REGION Network 9: Position Carrier Control First Carrier in Production Zone
   // Control of First Carrier in Zone Closest to end position/Stop.  Move command is issued to carrier. Carrier will move in auto.
   Label( ProdZoneFirstCarrierPosition )
   RUNG wire#powerrail
      Move(in := "EMS".Zone[#Zone].EndPos, out1 => #TrafficCopCarrierZnBufferOut[#CarrierZnArrayPos].CommandPos)
      Sub(in1 := #TrafficCopCarrierZnBufferOut[#CarrierZnArrayPos].CommandPos, in2 := "EMS".Zone[#Zone].InPositionTolerance, out => #TrafficCopCarrierZnBufferOut[#CarrierZnArrayPos].CommandPosLowLimit)
      Add(in1 := #TrafficCopCarrierZnBufferOut[#CarrierZnArrayPos].CommandPos, in2 := "EMS".Zone[#Zone].InPositionTolerance, out => #TrafficCopCarrierZnBufferOut[#CarrierZnArrayPos].CommandPosHighLimit)
   END_RUNG
   RUNG wire#powerrail
      { S7_Templates := "SrcType := DInt" } GE_Contact(in1 := "EMS".Carrier[#CarNumZnPos[1]].Position, in2 := #TrafficCopCarrierZnBufferOut[#CarrierZnArrayPos].CommandPosLowLimit)
      { S7_Templates := "SrcType := DInt" } LE_Contact(in1 := "EMS".Zone[#Zone].EndPos, in2 := #TrafficCopCarrierZnBufferOut[#CarrierZnArrayPos].CommandPosHighLimit)
      Coil( #TrafficCopCarrierZnBufferOut[#CarrierZnArrayPos].AtCommandPos )
   END_RUNG
   RUNG wire#powerrail
      Contact( "EMS".Carrier[#CarNumZnPos[1]].SDC_IN.AutoMode )
      I_Contact( #TrafficCopCarrierZnBufferOut[#CarrierZnArrayPos].AtCommandPos )
      Coil( #TCZnPosnArray.Carrier[#CarNumZnPos[#CarrierZnArrayPos]].MoveFwd )
   END_RUNG
   // the same network as SCL:
   ProdZoneFirstCarrierPosition:
   #TrafficCopCarrierZnBufferOut[#CarrierZnArrayPos].CommandPos := "EMS".Zone[#Zone].EndPos;
   #TrafficCopCarrierZnBufferOut[#CarrierZnArrayPos].CommandPosLowLimit := #TrafficCopCarrierZnBufferOut[#CarrierZnArrayPos].CommandPos - "EMS".Zone[#Zone].InPositionTolerance;
   #TrafficCopCarrierZnBufferOut[#CarrierZnArrayPos].CommandPosHighLimit := #TrafficCopCarrierZnBufferOut[#CarrierZnArrayPos].CommandPos + "EMS".Zone[#Zone].InPositionTolerance;
   #TrafficCopCarrierZnBufferOut[#CarrierZnArrayPos].AtCommandPos := ("EMS".Carrier[#CarNumZnPos[1]].Position >= #TrafficCopCarrierZnBufferOut[#CarrierZnArrayPos].CommandPosLowLimit) AND ("EMS".Zone[#Zone].EndPos <= #TrafficCopCarrierZnBufferOut[#CarrierZnArrayPos].CommandPosHighLimit);
   #TCZnPosnArray.Carrier[#CarNumZnPos[#CarrierZnArrayPos]].MoveFwd := "EMS".Carrier[#CarNumZnPos[1]].SDC_IN.AutoMode AND NOT #TrafficCopCarrierZnBufferOut[#CarrierZnArrayPos].AtCommandPos;
END_REGION

REGION Network 10: Start of 2nd to last Carrier in Zone Carrier Control
   Label( ZoneNextCarrierPosition )
   RUNG wire#powerrail
      Contact( "EMS".Zone[#Zone].AccumZone )
      JumpCoil( AccumZoneNextCarrierPosition )
   END_RUNG
   // the same network as SCL:
   ZoneNextCarrierPosition:
   IF "EMS".Zone[#Zone].AccumZone THEN GOTO AccumZoneNextCarrierPosition; END_IF;
END_REGION

REGION Network 11: Jump to Production Zone 2nd to Last Carrier Position Carrier Control
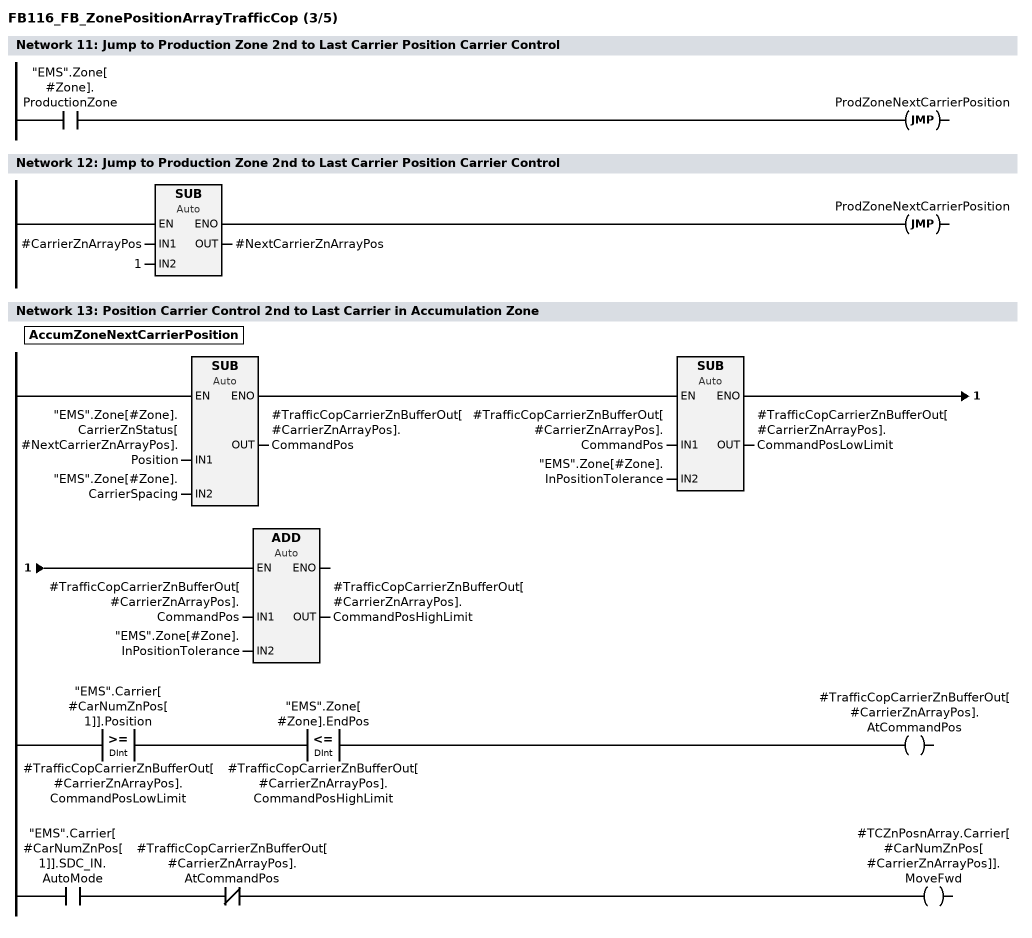
   RUNG wire#powerrail
      Contact( "EMS".Zone[#Zone].ProductionZone )
      JumpCoil( ProdZoneNextCarrierPosition )
   END_RUNG
   // the same network as SCL:
   IF "EMS".Zone[#Zone].ProductionZone THEN GOTO ProdZoneNextCarrierPosition; END_IF;
END_REGION

REGION Network 12: Jump to Production Zone 2nd to Last Carrier Position Carrier Control
   RUNG wire#powerrail
      Sub(in1 := #CarrierZnArrayPos, in2 := 1, out => #NextCarrierZnArrayPos)
      JumpCoil( ProdZoneNextCarrierPosition )
   END_RUNG
   // the same network as SCL:
   #NextCarrierZnArrayPos := #CarrierZnArrayPos - 1;
   GOTO ProdZoneNextCarrierPosition;
END_REGION

REGION Network 13: Position Carrier Control 2nd to Last Carrier in Accumulation Zone
   Label( AccumZoneNextCarrierPosition )
   RUNG wire#powerrail
      Sub(in1 := "EMS".Zone[#Zone].CarrierZnStatus[#NextCarrierZnArrayPos].Position, in2 := "EMS".Zone[#Zone].CarrierSpacing, out => #TrafficCopCarrierZnBufferOut[#CarrierZnArrayPos].CommandPos)
      Sub(in1 := #TrafficCopCarrierZnBufferOut[#CarrierZnArrayPos].CommandPos, in2 := "EMS".Zone[#Zone].InPositionTolerance, out => #TrafficCopCarrierZnBufferOut[#CarrierZnArrayPos].CommandPosLowLimit)
      Add(in1 := #TrafficCopCarrierZnBufferOut[#CarrierZnArrayPos].CommandPos, in2 := "EMS".Zone[#Zone].InPositionTolerance, out => #TrafficCopCarrierZnBufferOut[#CarrierZnArrayPos].CommandPosHighLimit)
   END_RUNG
   RUNG wire#powerrail
      { S7_Templates := "SrcType := DInt" } GE_Contact(in1 := "EMS".Carrier[#CarNumZnPos[1]].Position, in2 := #TrafficCopCarrierZnBufferOut[#CarrierZnArrayPos].CommandPosLowLimit)
      { S7_Templates := "SrcType := DInt" } LE_Contact(in1 := "EMS".Zone[#Zone].EndPos, in2 := #TrafficCopCarrierZnBufferOut[#CarrierZnArrayPos].CommandPosHighLimit)
      Coil( #TrafficCopCarrierZnBufferOut[#CarrierZnArrayPos].AtCommandPos )
   END_RUNG
   RUNG wire#powerrail
      Contact( "EMS".Carrier[#CarNumZnPos[1]].SDC_IN.AutoMode )
      I_Contact( #TrafficCopCarrierZnBufferOut[#CarrierZnArrayPos].AtCommandPos )
      Coil( #TCZnPosnArray.Carrier[#CarNumZnPos[#CarrierZnArrayPos]].MoveFwd )
   END_RUNG
   // the same network as SCL:
   AccumZoneNextCarrierPosition:
   #TrafficCopCarrierZnBufferOut[#CarrierZnArrayPos].CommandPos := "EMS".Zone[#Zone].CarrierZnStatus[#NextCarrierZnArrayPos].Position - "EMS".Zone[#Zone].CarrierSpacing;
   #TrafficCopCarrierZnBufferOut[#CarrierZnArrayPos].CommandPosLowLimit := #TrafficCopCarrierZnBufferOut[#CarrierZnArrayPos].CommandPos - "EMS".Zone[#Zone].InPositionTolerance;
   #TrafficCopCarrierZnBufferOut[#CarrierZnArrayPos].CommandPosHighLimit := #TrafficCopCarrierZnBufferOut[#CarrierZnArrayPos].CommandPos + "EMS".Zone[#Zone].InPositionTolerance;
   #TrafficCopCarrierZnBufferOut[#CarrierZnArrayPos].AtCommandPos := ("EMS".Carrier[#CarNumZnPos[1]].Position >= #TrafficCopCarrierZnBufferOut[#CarrierZnArrayPos].CommandPosLowLimit) AND ("EMS".Zone[#Zone].EndPos <= #TrafficCopCarrierZnBufferOut[#CarrierZnArrayPos].CommandPosHighLimit);
   #TCZnPosnArray.Carrier[#CarNumZnPos[#CarrierZnArrayPos]].MoveFwd := "EMS".Carrier[#CarNumZnPos[1]].SDC_IN.AutoMode AND NOT #TrafficCopCarrierZnBufferOut[#CarrierZnArrayPos].AtCommandPos;
END_REGION

REGION Network 14: Position Carrier Control 2nd to Last Carrier in Production Zone
   // Control of 2nd to Last Carrier in Zone Move to next zone with carrier spacing
   // .  Move command is issued to carrier. Carrier will move in auto.
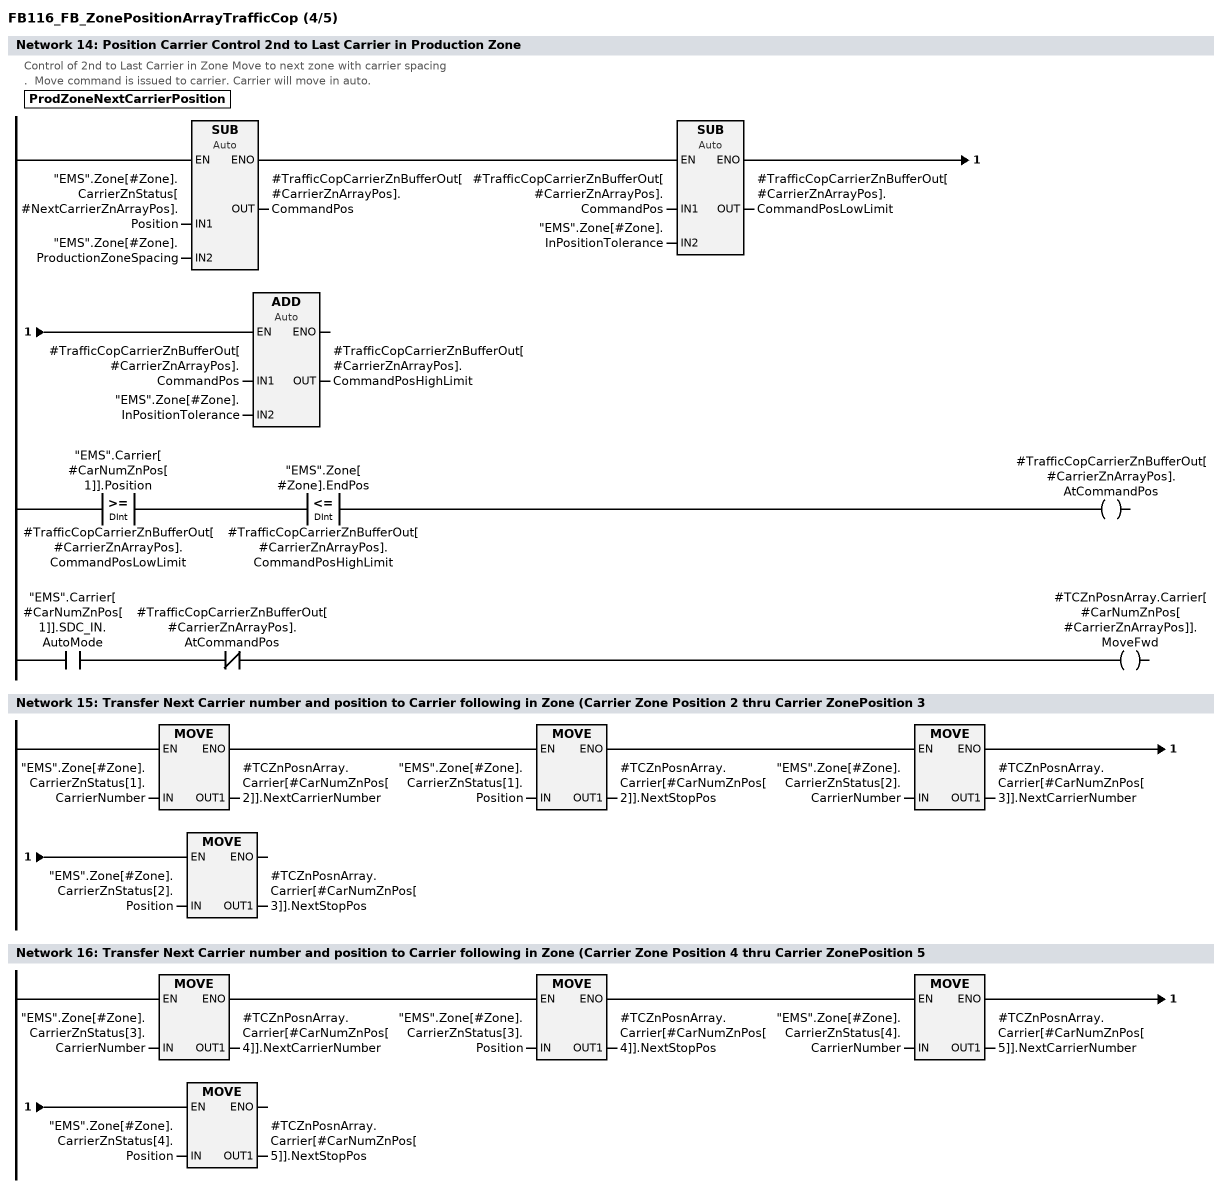
   Label( ProdZoneNextCarrierPosition )
   RUNG wire#powerrail
      Sub(in1 := "EMS".Zone[#Zone].CarrierZnStatus[#NextCarrierZnArrayPos].Position, in2 := "EMS".Zone[#Zone].ProductionZoneSpacing, out => #TrafficCopCarrierZnBufferOut[#CarrierZnArrayPos].CommandPos)
      Sub(in1 := #TrafficCopCarrierZnBufferOut[#CarrierZnArrayPos].CommandPos, in2 := "EMS".Zone[#Zone].InPositionTolerance, out => #TrafficCopCarrierZnBufferOut[#CarrierZnArrayPos].CommandPosLowLimit)
      Add(in1 := #TrafficCopCarrierZnBufferOut[#CarrierZnArrayPos].CommandPos, in2 := "EMS".Zone[#Zone].InPositionTolerance, out => #TrafficCopCarrierZnBufferOut[#CarrierZnArrayPos].CommandPosHighLimit)
   END_RUNG
   RUNG wire#powerrail
      { S7_Templates := "SrcType := DInt" } GE_Contact(in1 := "EMS".Carrier[#CarNumZnPos[1]].Position, in2 := #TrafficCopCarrierZnBufferOut[#CarrierZnArrayPos].CommandPosLowLimit)
      { S7_Templates := "SrcType := DInt" } LE_Contact(in1 := "EMS".Zone[#Zone].EndPos, in2 := #TrafficCopCarrierZnBufferOut[#CarrierZnArrayPos].CommandPosHighLimit)
      Coil( #TrafficCopCarrierZnBufferOut[#CarrierZnArrayPos].AtCommandPos )
   END_RUNG
   RUNG wire#powerrail
      Contact( "EMS".Carrier[#CarNumZnPos[1]].SDC_IN.AutoMode )
      I_Contact( #TrafficCopCarrierZnBufferOut[#CarrierZnArrayPos].AtCommandPos )
      Coil( #TCZnPosnArray.Carrier[#CarNumZnPos[#CarrierZnArrayPos]].MoveFwd )
   END_RUNG
   // the same network as SCL:
   ProdZoneNextCarrierPosition:
   #TrafficCopCarrierZnBufferOut[#CarrierZnArrayPos].CommandPos := "EMS".Zone[#Zone].CarrierZnStatus[#NextCarrierZnArrayPos].Position - "EMS".Zone[#Zone].ProductionZoneSpacing;
   #TrafficCopCarrierZnBufferOut[#CarrierZnArrayPos].CommandPosLowLimit := #TrafficCopCarrierZnBufferOut[#CarrierZnArrayPos].CommandPos - "EMS".Zone[#Zone].InPositionTolerance;
   #TrafficCopCarrierZnBufferOut[#CarrierZnArrayPos].CommandPosHighLimit := #TrafficCopCarrierZnBufferOut[#CarrierZnArrayPos].CommandPos + "EMS".Zone[#Zone].InPositionTolerance;
   #TrafficCopCarrierZnBufferOut[#CarrierZnArrayPos].AtCommandPos := ("EMS".Carrier[#CarNumZnPos[1]].Position >= #TrafficCopCarrierZnBufferOut[#CarrierZnArrayPos].CommandPosLowLimit) AND ("EMS".Zone[#Zone].EndPos <= #TrafficCopCarrierZnBufferOut[#CarrierZnArrayPos].CommandPosHighLimit);
   #TCZnPosnArray.Carrier[#CarNumZnPos[#CarrierZnArrayPos]].MoveFwd := "EMS".Carrier[#CarNumZnPos[1]].SDC_IN.AutoMode AND NOT #TrafficCopCarrierZnBufferOut[#CarrierZnArrayPos].AtCommandPos;
END_REGION

REGION Network 15: Transfer Next Carrier number and position to Carrier following in Zone (Carrier Zone Position 2 thru Carrier ZonePosition 3
   RUNG wire#powerrail
      Move(in := "EMS".Zone[#Zone].CarrierZnStatus[1].CarrierNumber, out1 => #TCZnPosnArray.Carrier[#CarNumZnPos[2]].NextCarrierNumber)
      Move(in := "EMS".Zone[#Zone].CarrierZnStatus[1].Position, out1 => #TCZnPosnArray.Carrier[#CarNumZnPos[2]].NextStopPos)
      Move(in := "EMS".Zone[#Zone].CarrierZnStatus[2].CarrierNumber, out1 => #TCZnPosnArray.Carrier[#CarNumZnPos[3]].NextCarrierNumber)
      Move(in := "EMS".Zone[#Zone].CarrierZnStatus[2].Position, out1 => #TCZnPosnArray.Carrier[#CarNumZnPos[3]].NextStopPos)
   END_RUNG
   // the same network as SCL:
   #TCZnPosnArray.Carrier[#CarNumZnPos[2]].NextCarrierNumber := "EMS".Zone[#Zone].CarrierZnStatus[1].CarrierNumber;
   #TCZnPosnArray.Carrier[#CarNumZnPos[2]].NextStopPos := "EMS".Zone[#Zone].CarrierZnStatus[1].Position;
   #TCZnPosnArray.Carrier[#CarNumZnPos[3]].NextCarrierNumber := "EMS".Zone[#Zone].CarrierZnStatus[2].CarrierNumber;
   #TCZnPosnArray.Carrier[#CarNumZnPos[3]].NextStopPos := "EMS".Zone[#Zone].CarrierZnStatus[2].Position;
END_REGION

REGION Network 16: Transfer Next Carrier number and position to Carrier following in Zone (Carrier Zone Position 4 thru Carrier ZonePosition 5
   RUNG wire#powerrail
      Move(in := "EMS".Zone[#Zone].CarrierZnStatus[3].CarrierNumber, out1 => #TCZnPosnArray.Carrier[#CarNumZnPos[4]].NextCarrierNumber)
      Move(in := "EMS".Zone[#Zone].CarrierZnStatus[3].Position, out1 => #TCZnPosnArray.Carrier[#CarNumZnPos[4]].NextStopPos)
      Move(in := "EMS".Zone[#Zone].CarrierZnStatus[4].CarrierNumber, out1 => #TCZnPosnArray.Carrier[#CarNumZnPos[5]].NextCarrierNumber)
      Move(in := "EMS".Zone[#Zone].CarrierZnStatus[4].Position, out1 => #TCZnPosnArray.Carrier[#CarNumZnPos[5]].NextStopPos)
   END_RUNG
   // the same network as SCL:
   #TCZnPosnArray.Carrier[#CarNumZnPos[4]].NextCarrierNumber := "EMS".Zone[#Zone].CarrierZnStatus[3].CarrierNumber;
   #TCZnPosnArray.Carrier[#CarNumZnPos[4]].NextStopPos := "EMS".Zone[#Zone].CarrierZnStatus[3].Position;
   #TCZnPosnArray.Carrier[#CarNumZnPos[5]].NextCarrierNumber := "EMS".Zone[#Zone].CarrierZnStatus[4].CarrierNumber;
   #TCZnPosnArray.Carrier[#CarNumZnPos[5]].NextStopPos := "EMS".Zone[#Zone].CarrierZnStatus[4].Position;
END_REGION

REGION Network 17: Transfer Next Carrier number and position to Carrier following in Zone (Carrier Zone Position 6 thru Carrier ZonePosition 7
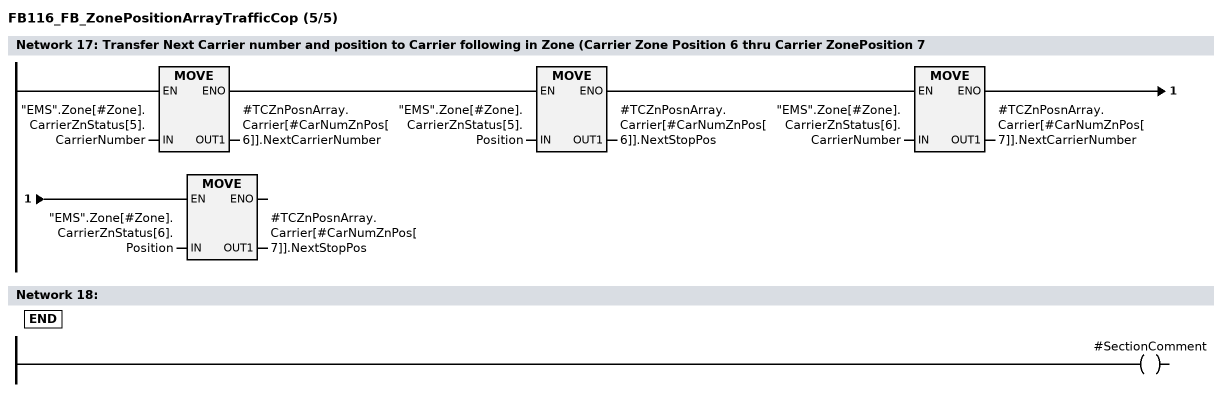
   RUNG wire#powerrail
      Move(in := "EMS".Zone[#Zone].CarrierZnStatus[5].CarrierNumber, out1 => #TCZnPosnArray.Carrier[#CarNumZnPos[6]].NextCarrierNumber)
      Move(in := "EMS".Zone[#Zone].CarrierZnStatus[5].Position, out1 => #TCZnPosnArray.Carrier[#CarNumZnPos[6]].NextStopPos)
      Move(in := "EMS".Zone[#Zone].CarrierZnStatus[6].CarrierNumber, out1 => #TCZnPosnArray.Carrier[#CarNumZnPos[7]].NextCarrierNumber)
      Move(in := "EMS".Zone[#Zone].CarrierZnStatus[6].Position, out1 => #TCZnPosnArray.Carrier[#CarNumZnPos[7]].NextStopPos)
   END_RUNG
   // the same network as SCL:
   #TCZnPosnArray.Carrier[#CarNumZnPos[6]].NextCarrierNumber := "EMS".Zone[#Zone].CarrierZnStatus[5].CarrierNumber;
   #TCZnPosnArray.Carrier[#CarNumZnPos[6]].NextStopPos := "EMS".Zone[#Zone].CarrierZnStatus[5].Position;
   #TCZnPosnArray.Carrier[#CarNumZnPos[7]].NextCarrierNumber := "EMS".Zone[#Zone].CarrierZnStatus[6].CarrierNumber;
   #TCZnPosnArray.Carrier[#CarNumZnPos[7]].NextStopPos := "EMS".Zone[#Zone].CarrierZnStatus[6].Position;
END_REGION

REGION Network 18
   Label( END )
   RUNG wire#powerrail
      Coil( #SectionComment )
   END_RUNG
   // the same network as SCL:
   END:
   #SectionComment := TRUE;
END_REGION
END_FUNCTION_BLOCK

FUNCTION_BLOCK "FB117_MapSDCOut_Carrier"   // FB117, LAD
{ S7_Optimized_Access := 'TRUE' }
VERSION : 0.1
   VAR_INPUT
      ZoneArray : Array[0..60] of "UDT_TC_SDCOutZone";
      Carrier : Int;
      Zone : Int;
   END_VAR
   VAR_OUTPUT
      DriveFwdCMD : Bool;
      AtCmdPos : Bool;
      NextStopPos : DWord;
      DriveCmdSpeed : Int;
      Zone_Echo : Int;
      Pos_Echo : DWord;
   END_VAR
   VAR
      CarrierArray : Array[0..99] of "UDT_TC_SDCOutCarrier";
   END_VAR
   VAR_TEMP   // added for the SCL form of the ladder/FBD networks
      _w1 : Bool;
   END_VAR
BEGIN

REGION Network 1
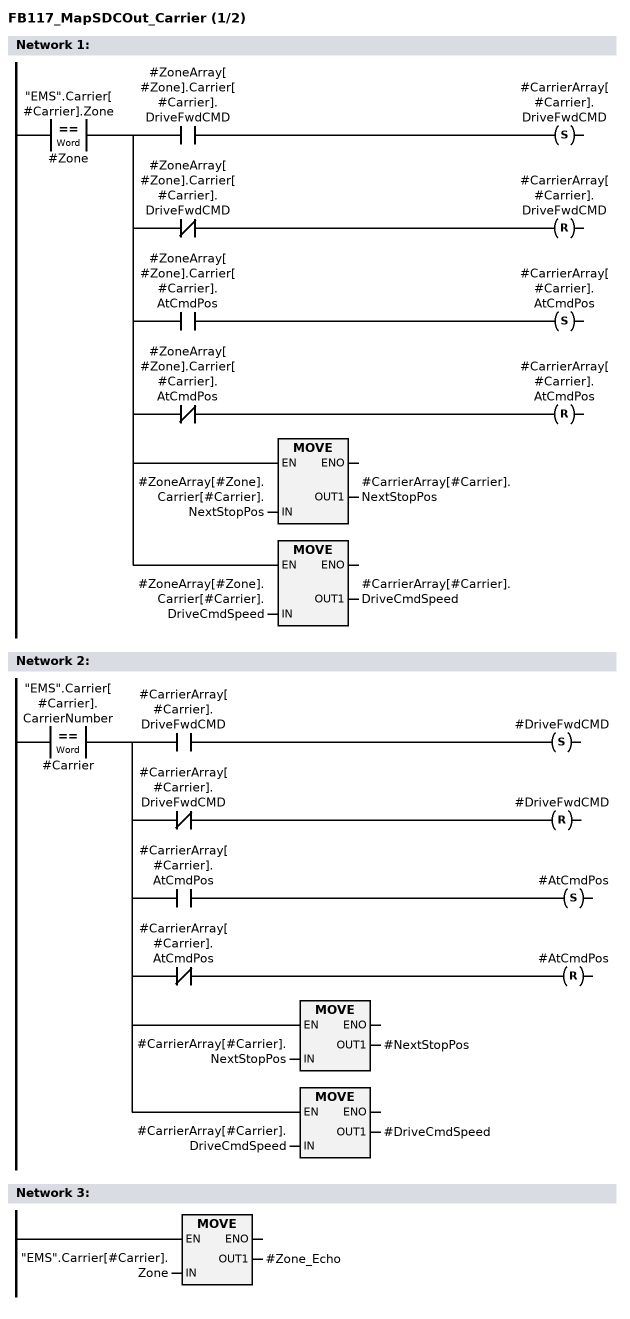
   RUNG wire#powerrail
      { S7_Templates := "SrcType := Word" } EQ_Contact(in1 := "EMS".Carrier[#Carrier].Zone, in2 := #Zone)
      wire#w1
      Contact( #ZoneArray[#Zone].Carrier[#Carrier].DriveFwdCMD )
      S_Coil( #CarrierArray[#Carrier].DriveFwdCMD )
   END_RUNG
   RUNG wire#w1
      I_Contact( #ZoneArray[#Zone].Carrier[#Carrier].DriveFwdCMD )
      R_Coil( #CarrierArray[#Carrier].DriveFwdCMD )
   END_RUNG
   RUNG wire#w1
      Contact( #ZoneArray[#Zone].Carrier[#Carrier].AtCmdPos )
      S_Coil( #CarrierArray[#Carrier].AtCmdPos )
   END_RUNG
   RUNG wire#w1
      I_Contact( #ZoneArray[#Zone].Carrier[#Carrier].AtCmdPos )
      R_Coil( #CarrierArray[#Carrier].AtCmdPos )
   END_RUNG
   RUNG wire#w1
      Move(in := #ZoneArray[#Zone].Carrier[#Carrier].NextStopPos, out1 => #CarrierArray[#Carrier].NextStopPos)
   END_RUNG
   RUNG wire#w1
      Move(in := #ZoneArray[#Zone].Carrier[#Carrier].DriveCmdSpeed, out1 => #CarrierArray[#Carrier].DriveCmdSpeed)
   END_RUNG
   // the same network as SCL:
   #_w1 := "EMS".Carrier[#Carrier].Zone = #Zone;
   IF #_w1 AND #ZoneArray[#Zone].Carrier[#Carrier].DriveFwdCMD THEN
       #CarrierArray[#Carrier].DriveFwdCMD := TRUE;
   END_IF;
   IF #_w1 AND NOT #ZoneArray[#Zone].Carrier[#Carrier].DriveFwdCMD THEN
       #CarrierArray[#Carrier].DriveFwdCMD := FALSE;
   END_IF;
   IF #_w1 AND #ZoneArray[#Zone].Carrier[#Carrier].AtCmdPos THEN
       #CarrierArray[#Carrier].AtCmdPos := TRUE;
   END_IF;
   IF #_w1 AND NOT #ZoneArray[#Zone].Carrier[#Carrier].AtCmdPos THEN
       #CarrierArray[#Carrier].AtCmdPos := FALSE;
   END_IF;
   IF #_w1 THEN
       #CarrierArray[#Carrier].NextStopPos := #ZoneArray[#Zone].Carrier[#Carrier].NextStopPos;
       #CarrierArray[#Carrier].DriveCmdSpeed := #ZoneArray[#Zone].Carrier[#Carrier].DriveCmdSpeed;
   END_IF;
END_REGION

REGION Network 2
   RUNG wire#powerrail
      { S7_Templates := "SrcType := Word" } EQ_Contact(in1 := "EMS".Carrier[#Carrier].CarrierNumber, in2 := #Carrier)
      wire#w1
      Contact( #CarrierArray[#Carrier].DriveFwdCMD )
      S_Coil( #DriveFwdCMD )
   END_RUNG
   RUNG wire#w1
      I_Contact( #CarrierArray[#Carrier].DriveFwdCMD )
      R_Coil( #DriveFwdCMD )
   END_RUNG
   RUNG wire#w1
      Contact( #CarrierArray[#Carrier].AtCmdPos )
      S_Coil( #AtCmdPos )
   END_RUNG
   RUNG wire#w1
      I_Contact( #CarrierArray[#Carrier].AtCmdPos )
      R_Coil( #AtCmdPos )
   END_RUNG
   RUNG wire#w1
      Move(in := #CarrierArray[#Carrier].NextStopPos, out1 => #NextStopPos)
   END_RUNG
   RUNG wire#w1
      Move(in := #CarrierArray[#Carrier].DriveCmdSpeed, out1 => #DriveCmdSpeed)
   END_RUNG
   // the same network as SCL:
   #_w1 := "EMS".Carrier[#Carrier].CarrierNumber = #Carrier;
   IF #_w1 AND #CarrierArray[#Carrier].DriveFwdCMD THEN #DriveFwdCMD := TRUE; END_IF;
   IF #_w1 AND NOT #CarrierArray[#Carrier].DriveFwdCMD THEN #DriveFwdCMD := FALSE; END_IF;
   IF #_w1 AND #CarrierArray[#Carrier].AtCmdPos THEN #AtCmdPos := TRUE; END_IF;
   IF #_w1 AND NOT #CarrierArray[#Carrier].AtCmdPos THEN #AtCmdPos := FALSE; END_IF;
   IF #_w1 THEN
       #NextStopPos := #CarrierArray[#Carrier].NextStopPos;
       #DriveCmdSpeed := #CarrierArray[#Carrier].DriveCmdSpeed;
   END_IF;
END_REGION

REGION Network 3
   RUNG wire#powerrail
      Move(in := "EMS".Carrier[#Carrier].Zone, out1 => #Zone_Echo)
   END_RUNG
   // the same network as SCL:
   #Zone_Echo := "EMS".Carrier[#Carrier].Zone;
END_REGION

REGION Network 4
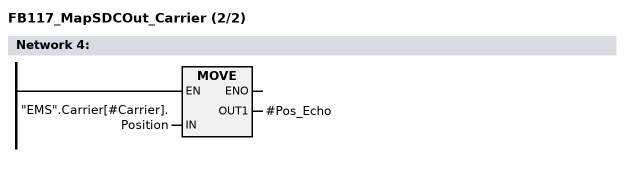
   RUNG wire#powerrail
      Move(in := "EMS".Carrier[#Carrier].Position, out1 => #Pos_Echo)
   END_RUNG
   // the same network as SCL:
   #Pos_Echo := "EMS".Carrier[#Carrier].Position;
END_REGION
END_FUNCTION_BLOCK

FUNCTION_BLOCK "FB118_TCMapSDCOut"   // FB118, LAD
{ S7_Optimized_Access := 'TRUE' }
VERSION : 0.1
   VAR_INPUT
      TC_ZoneMotion : "UDT_TC_ZoneMotion";
      Zone : Int;
      Carrier : Int;
   END_VAR
   VAR_OUTPUT
      SDC_Out : Array[0..99] of "UDT_SDC_OUT";
      SDCOUT_DriveFwdCmd : Bool;
      SDCOUT_DriveCmdSpeed : Word;
      SDCOUT_NextStopPos : DWord;
      SDCOUT_NextCarrierNum : Word;
      SDCOut_AtCmdPos : Bool;
   END_VAR
   VAR
      CarrierTempZone : Int;
      oneshot : Array[0..20] of Bool;
      oneshotneg : Bool;
      oneshot3 : Bool;
      resetlatch1 : Bool;
      DriveCmdSetup : Array[0..99] of Bool;
   END_VAR
   VAR_TEMP
      tempptrig : Bool;
   END_VAR
BEGIN

REGION Network 1
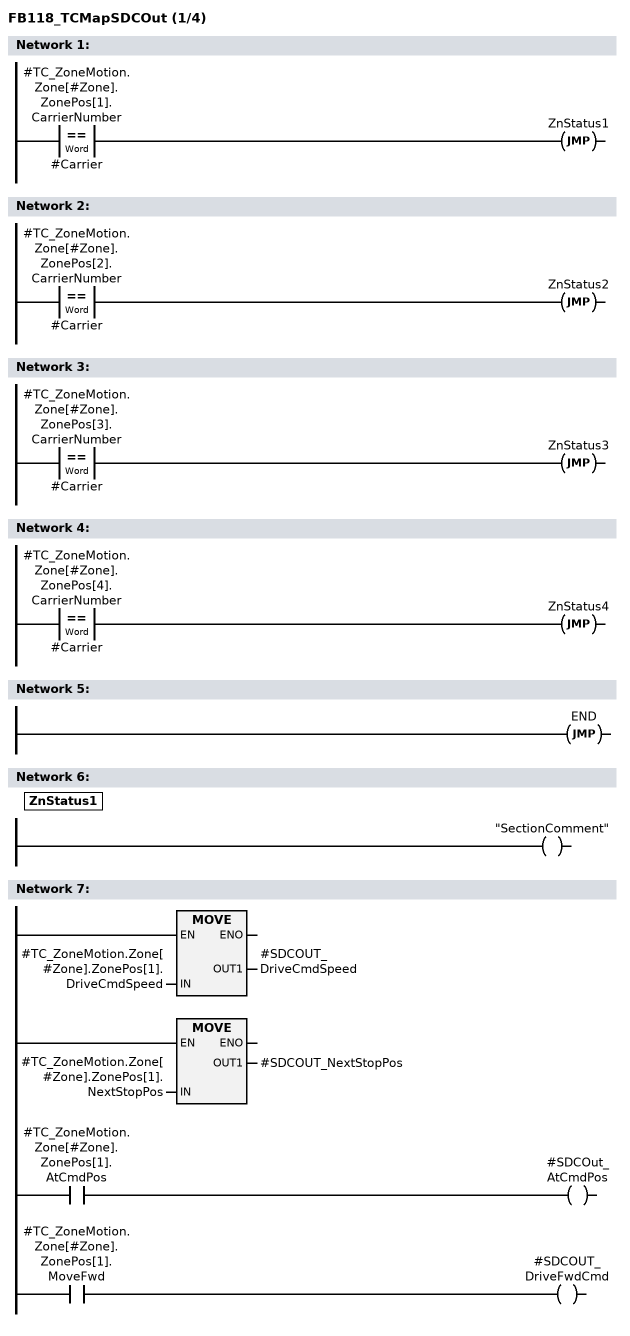
   RUNG wire#powerrail
      { S7_Templates := "SrcType := Word" } EQ_Contact(in1 := #TC_ZoneMotion.Zone[#Zone].ZonePos[1].CarrierNumber, in2 := #Carrier)
      JumpCoil( ZnStatus1 )
   END_RUNG
   // the same network as SCL:
   IF #TC_ZoneMotion.Zone[#Zone].ZonePos[1].CarrierNumber = #Carrier THEN GOTO ZnStatus1; END_IF;
END_REGION

REGION Network 2
   RUNG wire#powerrail
      { S7_Templates := "SrcType := Word" } EQ_Contact(in1 := #TC_ZoneMotion.Zone[#Zone].ZonePos[2].CarrierNumber, in2 := #Carrier)
      JumpCoil( ZnStatus2 )
   END_RUNG
   // the same network as SCL:
   IF #TC_ZoneMotion.Zone[#Zone].ZonePos[2].CarrierNumber = #Carrier THEN GOTO ZnStatus2; END_IF;
END_REGION

REGION Network 3
   RUNG wire#powerrail
      { S7_Templates := "SrcType := Word" } EQ_Contact(in1 := #TC_ZoneMotion.Zone[#Zone].ZonePos[3].CarrierNumber, in2 := #Carrier)
      JumpCoil( ZnStatus3 )
   END_RUNG
   // the same network as SCL:
   IF #TC_ZoneMotion.Zone[#Zone].ZonePos[3].CarrierNumber = #Carrier THEN GOTO ZnStatus3; END_IF;
END_REGION

REGION Network 4
   RUNG wire#powerrail
      { S7_Templates := "SrcType := Word" } EQ_Contact(in1 := #TC_ZoneMotion.Zone[#Zone].ZonePos[4].CarrierNumber, in2 := #Carrier)
      JumpCoil( ZnStatus4 )
   END_RUNG
   // the same network as SCL:
   IF #TC_ZoneMotion.Zone[#Zone].ZonePos[4].CarrierNumber = #Carrier THEN GOTO ZnStatus4; END_IF;
END_REGION

REGION Network 5
   RUNG wire#powerrail
      JumpCoil( END )
   END_RUNG
   // the same network as SCL:
   GOTO END;
END_REGION

REGION Network 6
   Label( ZnStatus1 )
   RUNG wire#powerrail
      Coil( "SectionComment" )
   END_RUNG
   // the same network as SCL:
   ZnStatus1:
   "SectionComment" := TRUE;
END_REGION

REGION Network 7
   RUNG wire#powerrail
      Move(in := #TC_ZoneMotion.Zone[#Zone].ZonePos[1].DriveCmdSpeed, out1 => #SDCOUT_DriveCmdSpeed)
   END_RUNG
   RUNG wire#powerrail
      Move(in := #TC_ZoneMotion.Zone[#Zone].ZonePos[1].NextStopPos, out1 => #SDCOUT_NextStopPos)
   END_RUNG
   RUNG wire#powerrail
      Contact( #TC_ZoneMotion.Zone[#Zone].ZonePos[1].AtCmdPos )
      Coil( #SDCOut_AtCmdPos )
   END_RUNG
   RUNG wire#powerrail
      Contact( #TC_ZoneMotion.Zone[#Zone].ZonePos[1].MoveFwd )
      Coil( #SDCOUT_DriveFwdCmd )
   END_RUNG
   // the same network as SCL:
   #SDCOUT_DriveCmdSpeed := #TC_ZoneMotion.Zone[#Zone].ZonePos[1].DriveCmdSpeed;
   #SDCOUT_NextStopPos := #TC_ZoneMotion.Zone[#Zone].ZonePos[1].NextStopPos;
   #SDCOut_AtCmdPos := #TC_ZoneMotion.Zone[#Zone].ZonePos[1].AtCmdPos;
   #SDCOUT_DriveFwdCmd := #TC_ZoneMotion.Zone[#Zone].ZonePos[1].MoveFwd;
END_REGION

REGION Network 8
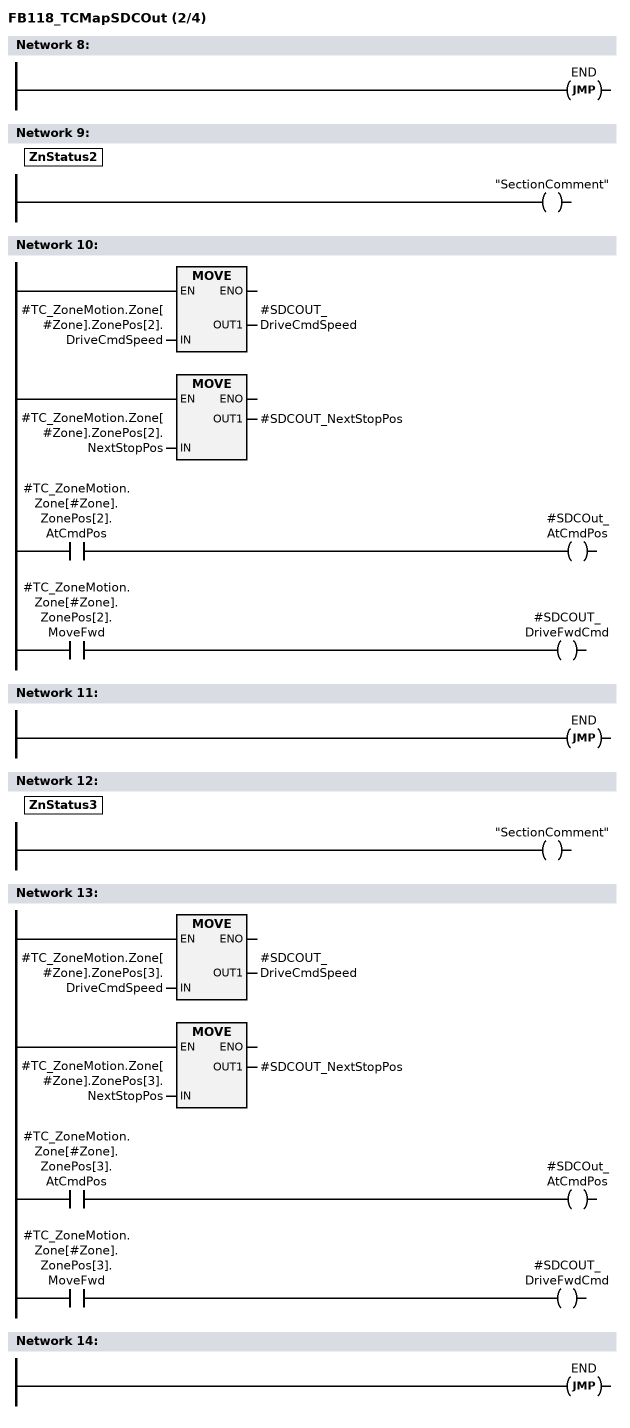
   RUNG wire#powerrail
      JumpCoil( END )
   END_RUNG
   // the same network as SCL:
   GOTO END;
END_REGION

REGION Network 9
   Label( ZnStatus2 )
   RUNG wire#powerrail
      Coil( "SectionComment" )
   END_RUNG
   // the same network as SCL:
   ZnStatus2:
   "SectionComment" := TRUE;
END_REGION

REGION Network 10
   RUNG wire#powerrail
      Move(in := #TC_ZoneMotion.Zone[#Zone].ZonePos[2].DriveCmdSpeed, out1 => #SDCOUT_DriveCmdSpeed)
   END_RUNG
   RUNG wire#powerrail
      Move(in := #TC_ZoneMotion.Zone[#Zone].ZonePos[2].NextStopPos, out1 => #SDCOUT_NextStopPos)
   END_RUNG
   RUNG wire#powerrail
      Contact( #TC_ZoneMotion.Zone[#Zone].ZonePos[2].AtCmdPos )
      Coil( #SDCOut_AtCmdPos )
   END_RUNG
   RUNG wire#powerrail
      Contact( #TC_ZoneMotion.Zone[#Zone].ZonePos[2].MoveFwd )
      Coil( #SDCOUT_DriveFwdCmd )
   END_RUNG
   // the same network as SCL:
   #SDCOUT_DriveCmdSpeed := #TC_ZoneMotion.Zone[#Zone].ZonePos[2].DriveCmdSpeed;
   #SDCOUT_NextStopPos := #TC_ZoneMotion.Zone[#Zone].ZonePos[2].NextStopPos;
   #SDCOut_AtCmdPos := #TC_ZoneMotion.Zone[#Zone].ZonePos[2].AtCmdPos;
   #SDCOUT_DriveFwdCmd := #TC_ZoneMotion.Zone[#Zone].ZonePos[2].MoveFwd;
END_REGION

REGION Network 11
   RUNG wire#powerrail
      JumpCoil( END )
   END_RUNG
   // the same network as SCL:
   GOTO END;
END_REGION

REGION Network 12
   Label( ZnStatus3 )
   RUNG wire#powerrail
      Coil( "SectionComment" )
   END_RUNG
   // the same network as SCL:
   ZnStatus3:
   "SectionComment" := TRUE;
END_REGION

REGION Network 13
   RUNG wire#powerrail
      Move(in := #TC_ZoneMotion.Zone[#Zone].ZonePos[3].DriveCmdSpeed, out1 => #SDCOUT_DriveCmdSpeed)
   END_RUNG
   RUNG wire#powerrail
      Move(in := #TC_ZoneMotion.Zone[#Zone].ZonePos[3].NextStopPos, out1 => #SDCOUT_NextStopPos)
   END_RUNG
   RUNG wire#powerrail
      Contact( #TC_ZoneMotion.Zone[#Zone].ZonePos[3].AtCmdPos )
      Coil( #SDCOut_AtCmdPos )
   END_RUNG
   RUNG wire#powerrail
      Contact( #TC_ZoneMotion.Zone[#Zone].ZonePos[3].MoveFwd )
      Coil( #SDCOUT_DriveFwdCmd )
   END_RUNG
   // the same network as SCL:
   #SDCOUT_DriveCmdSpeed := #TC_ZoneMotion.Zone[#Zone].ZonePos[3].DriveCmdSpeed;
   #SDCOUT_NextStopPos := #TC_ZoneMotion.Zone[#Zone].ZonePos[3].NextStopPos;
   #SDCOut_AtCmdPos := #TC_ZoneMotion.Zone[#Zone].ZonePos[3].AtCmdPos;
   #SDCOUT_DriveFwdCmd := #TC_ZoneMotion.Zone[#Zone].ZonePos[3].MoveFwd;
END_REGION

REGION Network 14
   RUNG wire#powerrail
      JumpCoil( END )
   END_RUNG
   // the same network as SCL:
   GOTO END;
END_REGION

REGION Network 15
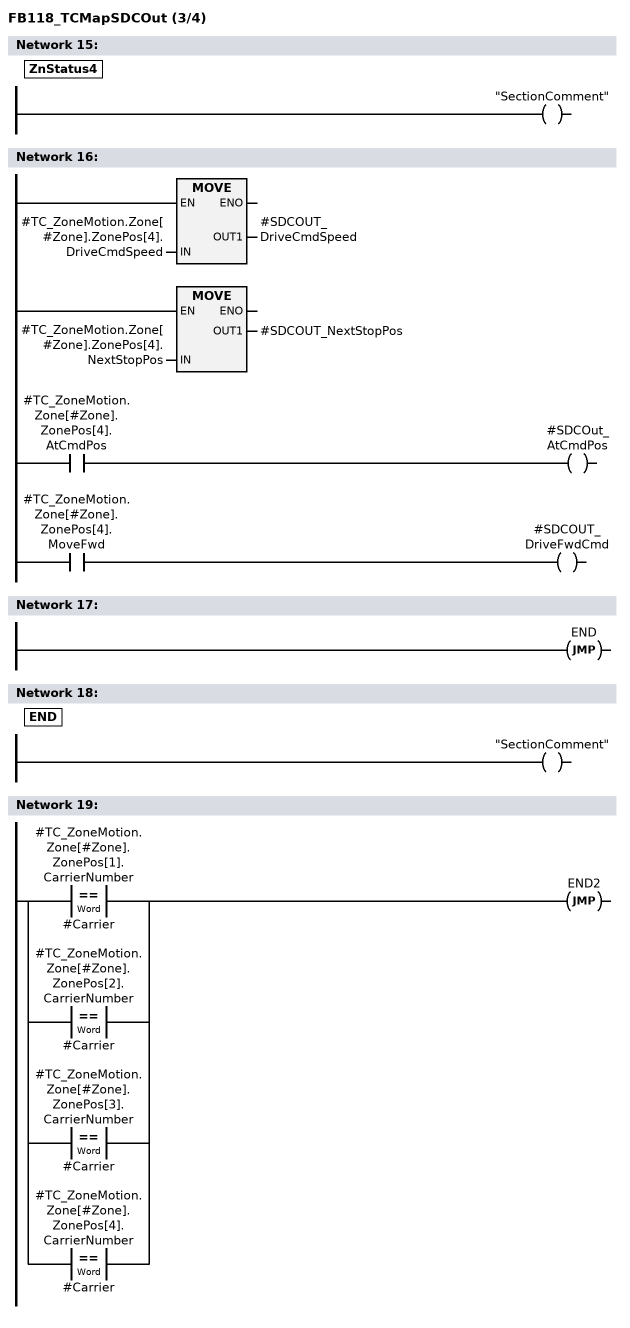
   Label( ZnStatus4 )
   RUNG wire#powerrail
      Coil( "SectionComment" )
   END_RUNG
   // the same network as SCL:
   ZnStatus4:
   "SectionComment" := TRUE;
END_REGION

REGION Network 16
   RUNG wire#powerrail
      Move(in := #TC_ZoneMotion.Zone[#Zone].ZonePos[4].DriveCmdSpeed, out1 => #SDCOUT_DriveCmdSpeed)
   END_RUNG
   RUNG wire#powerrail
      Move(in := #TC_ZoneMotion.Zone[#Zone].ZonePos[4].NextStopPos, out1 => #SDCOUT_NextStopPos)
   END_RUNG
   RUNG wire#powerrail
      Contact( #TC_ZoneMotion.Zone[#Zone].ZonePos[4].AtCmdPos )
      Coil( #SDCOut_AtCmdPos )
   END_RUNG
   RUNG wire#powerrail
      Contact( #TC_ZoneMotion.Zone[#Zone].ZonePos[4].MoveFwd )
      Coil( #SDCOUT_DriveFwdCmd )
   END_RUNG
   // the same network as SCL:
   #SDCOUT_DriveCmdSpeed := #TC_ZoneMotion.Zone[#Zone].ZonePos[4].DriveCmdSpeed;
   #SDCOUT_NextStopPos := #TC_ZoneMotion.Zone[#Zone].ZonePos[4].NextStopPos;
   #SDCOut_AtCmdPos := #TC_ZoneMotion.Zone[#Zone].ZonePos[4].AtCmdPos;
   #SDCOUT_DriveFwdCmd := #TC_ZoneMotion.Zone[#Zone].ZonePos[4].MoveFwd;
END_REGION

REGION Network 17
   RUNG wire#powerrail
      JumpCoil( END )
   END_RUNG
   // the same network as SCL:
   GOTO END;
END_REGION

REGION Network 18
   Label( END )
   RUNG wire#powerrail
      Coil( "SectionComment" )
   END_RUNG
   // the same network as SCL:
   END:
   "SectionComment" := TRUE;
END_REGION

REGION Network 19
   RUNG wire#powerrail
      { S7_Templates := "SrcType := Word" } EQ_Contact(in1 := #TC_ZoneMotion.Zone[#Zone].ZonePos[1].CarrierNumber, in2 := #Carrier)
      wire#w1
      JumpCoil( END2 )
   END_RUNG
   RUNG wire#powerrail
      { S7_Templates := "SrcType := Word" } EQ_Contact(in1 := #TC_ZoneMotion.Zone[#Zone].ZonePos[2].CarrierNumber, in2 := #Carrier)
   END_RUNG wire#w1
   RUNG wire#powerrail
      { S7_Templates := "SrcType := Word" } EQ_Contact(in1 := #TC_ZoneMotion.Zone[#Zone].ZonePos[3].CarrierNumber, in2 := #Carrier)
   END_RUNG wire#w1
   RUNG wire#powerrail
      { S7_Templates := "SrcType := Word" } EQ_Contact(in1 := #TC_ZoneMotion.Zone[#Zone].ZonePos[4].CarrierNumber, in2 := #Carrier)
   END_RUNG wire#w1
   // the same network as SCL:
   IF (#TC_ZoneMotion.Zone[#Zone].ZonePos[1].CarrierNumber = #Carrier) OR (#TC_ZoneMotion.Zone[#Zone].ZonePos[2].CarrierNumber = #Carrier) OR (#TC_ZoneMotion.Zone[#Zone].ZonePos[3].CarrierNumber = #Carrier) OR (#TC_ZoneMotion.Zone[#Zone].ZonePos[4].CarrierNumber = #Carrier) THEN
       GOTO END2;
   END_IF;
END_REGION

REGION Network 20
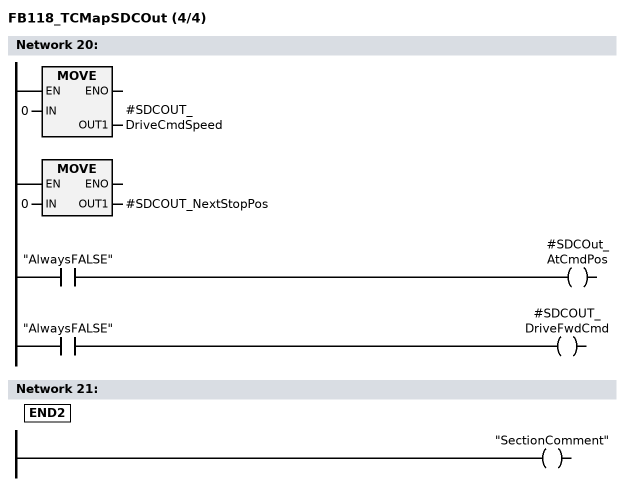
   RUNG wire#powerrail
      Move(in := 0, out1 => #SDCOUT_DriveCmdSpeed)
   END_RUNG
   RUNG wire#powerrail
      Move(in := 0, out1 => #SDCOUT_NextStopPos)
   END_RUNG
   RUNG wire#powerrail
      Contact( "AlwaysFALSE" )
      Coil( #SDCOut_AtCmdPos )
   END_RUNG
   RUNG wire#powerrail
      Contact( "AlwaysFALSE" )
      Coil( #SDCOUT_DriveFwdCmd )
   END_RUNG
   // the same network as SCL:
   #SDCOUT_DriveCmdSpeed := 0;
   #SDCOUT_NextStopPos := 0;
   #SDCOut_AtCmdPos := "AlwaysFALSE";
   #SDCOUT_DriveFwdCmd := "AlwaysFALSE";
END_REGION

REGION Network 21
   Label( END2 )
   RUNG wire#powerrail
      Coil( "SectionComment" )
   END_RUNG
   // the same network as SCL:
   END2:
   "SectionComment" := TRUE;
END_REGION
END_FUNCTION_BLOCK

FUNCTION_BLOCK "FB119_ZoneTrafficCop"   // FB119, LAD
{ S7_Optimized_Access := 'FALSE' }
VERSION : 0.1
   VAR_INPUT
      EMS : "UDT_System";
      Zone : Int := 1;
   END_VAR
   VAR_OUTPUT
      TrafficCopZone : "UDT_TrafficCopZoneStructure";
   END_VAR
   VAR
      SectionComment : Bool;
      TotalZonePositions : Int;
   END_VAR
BEGIN

REGION Network 1: Section Comment
   // Section Logic for Current Carrier number in Position 1 - Max Carrier in Zone Position Array
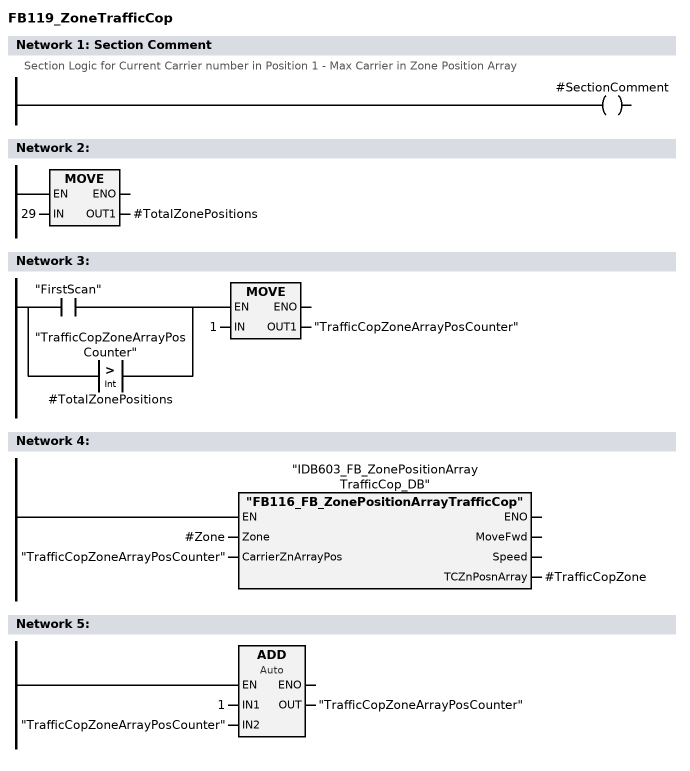
   RUNG wire#powerrail
      Coil( #SectionComment )
   END_RUNG
   // the same network as SCL:
   #SectionComment := TRUE;
END_REGION

REGION Network 2
   RUNG wire#powerrail
      Move(in := 29, out1 => #TotalZonePositions)
   END_RUNG
   // the same network as SCL:
   #TotalZonePositions := 29;
END_REGION

REGION Network 3
   RUNG wire#powerrail
      Contact( "FirstScan" )
      wire#w1
      Move(in := 1, out1 => "TrafficCopZoneArrayPosCounter")
   END_RUNG
   RUNG wire#powerrail
      { S7_Templates := "SrcType := Int" } GT_Contact(in1 := "TrafficCopZoneArrayPosCounter", in2 := #TotalZonePositions)
   END_RUNG wire#w1
   // the same network as SCL:
   IF "FirstScan" OR ("TrafficCopZoneArrayPosCounter" > #TotalZonePositions) THEN
       "TrafficCopZoneArrayPosCounter" := 1;
   END_IF;
END_REGION

REGION Network 4
   RUNG wire#powerrail
      "IDB603_FB_ZonePositionArrayTrafficCop_DB"(Zone := #Zone, CarrierZnArrayPos := "TrafficCopZoneArrayPosCounter", MoveFwd =>, Speed =>, TCZnPosnArray => #TrafficCopZone)
   END_RUNG
   // the same network as SCL:
   "IDB603_FB_ZonePositionArrayTrafficCop_DB"(Zone := #Zone,   // "FB116_FB_ZonePositionArrayTrafficCop"
                           CarrierZnArrayPos := "TrafficCopZoneArrayPosCounter",
                           TCZnPosnArray => #TrafficCopZone);
END_REGION

REGION Network 5
   RUNG wire#powerrail
      Add(in1 := 1, in2 := "TrafficCopZoneArrayPosCounter", out => "TrafficCopZoneArrayPosCounter")
   END_RUNG
   // the same network as SCL:
   "TrafficCopZoneArrayPosCounter" := 1 + "TrafficCopZoneArrayPosCounter";
END_REGION
END_FUNCTION_BLOCK

FUNCTION_BLOCK "FB120_ZoneSpacingCheck"   // FB120, SCL
{ S7_Optimized_Access := 'TRUE' }
VERSION : 0.1
   VAR_INPUT
      Zone : Int;
      TotalPosition : Int;
      EMS : "UDT_System";
   END_VAR
   VAR_OUTPUT
      GapSpacingFault : Bool;
      GapFaultZnPosition : Int;
      FirstCarrierNumGapFlt : Int;
      SecondCarrierNumGapFlt : Int;
   END_VAR
   VAR_TEMP
      ZnPosCounter : Int;
      ZoneFound : Word;
      FirstHighPos : Int;
      FirstLowPos : Int;
      NextLowPos : Int;
      NextHighPos : Int;
      GapSpaceActual : Int;
      GapSpaceActualhiLimit : Int;
      GapSpaceActualLowLimit : Int;
      NextZnPosCounter : Int;
      MaxGapSpacing : Int;
   END_VAR
BEGIN
       #ZnPosCounter := 1;
       #GapSpacingFault := 0;
       #GapFaultZnPosition := 0;
       #FirstCarrierNumGapFlt := 0;
       #SecondCarrierNumGapFlt := 0;
       FOR #ZnPosCounter := 1 TO #TotalPosition DO
           #NextZnPosCounter := #ZnPosCounter + 1;
           IF #EMS.Zone[#Zone].CarrierZnStatus[#NextZnPosCounter].CarrierNumber = 0 THEN
               ;
               RETURN;
           END_IF;

           #GapSpaceActual := #EMS.Zone[#Zone].CarrierZnStatus[#ZnPosCounter].Position - #EMS.Zone[#Zone].CarrierZnStatus[#NextZnPosCounter].Position;
           #MaxGapSpacing := #GapSpaceActual + #EMS.Zone[#Zone].InPositionTolerance;
           IF #EMS.Zone[#Zone].AccumZone = 1 & #MaxGapSpacing < #EMS.Zone[#Zone].CarrierSpacing OR #EMS.Zone[#Zone].ProductionZone = 1 & #MaxGapSpacing < #EMS.Zone[#Zone].ProductionZoneSpacing THEN
               #GapSpacingFault := 1;
               #GapFaultZnPosition := #ZnPosCounter;
               #FirstCarrierNumGapFlt := #EMS.Zone[#Zone].CarrierZnStatus[#ZnPosCounter].CarrierNumber;
               #SecondCarrierNumGapFlt := #EMS.Zone[#Zone].CarrierZnStatus[#NextZnPosCounter].CarrierNumber;
          ELSE
    #GapSpacingFault := 0;
     //#FirstCarrierNumGapFlt := 0;
     //#SecondCarrierNumGapFlt := 0;
               RETURN;
           END_IF;
       END_FOR;
END_FUNCTION_BLOCK

// folder: 04_FCs

FUNCTION "FC100_EMS_System" : Void   // FC100, LAD
{ S7_Optimized_Access := 'TRUE' }
VERSION : 0.1
   VAR_TEMP
      TEMPCARRIERNUMBR : Word;
   END_VAR
BEGIN

REGION Network 1